REGION Network 7: LS425, LS442 Alarms (RIO 07: APT)
   RUNG wire#powerrail
      "1602_DIGITAL_HEALTH"(InputSignal := "20_TANKS_IP_DATA".RIO_07.FIRST_TANK.BWT_LEVEL_HIHI, InputTripLevel := #InputTripLevel, SensorHealthOut => "1092_HMI_OP_FLAGS".LS425_442_LevelSwitch_HighHigh_Alarm[14].Healthy, AlarmOut => "1092_HMI_OP_FLAGS".LS425_442_LevelSwitch_HighHigh_Alarm[14].UnhealthyAlarm)
   END_RUNG
   // the same network as SCL:
   "1602_DIGITAL_HEALTH"(InputSignal := "20_TANKS_IP_DATA".RIO_07.FIRST_TANK.BWT_LEVEL_HIHI,
                         InputTripLevel := #InputTripLevel,
                         SensorHealthOut => "1092_HMI_OP_FLAGS".LS425_442_LevelSwitch_HighHigh_Alarm[14].Healthy,
                         AlarmOut => "1092_HMI_OP_FLAGS".LS425_442_LevelSwitch_HighHigh_Alarm[14].UnhealthyAlarm);
END_REGION
END_FUNCTION

// folder: 1000 - 1999 BWT System Control/1060 - 1089 Alarm & Valve Status Handling/1080 - 1084 Tank Group Alarms

FUNCTION "1080_PT424_ALARMS" : Void   // FC1080, LAD
{ S7_Optimized_Access := 'TRUE' }
VERSION : 0.1
// Alarm wrapper function for Ullage Space Pressure Transmitter on each tank group.
BEGIN

REGION Network 1: PT424 Alarms (RIO 01)
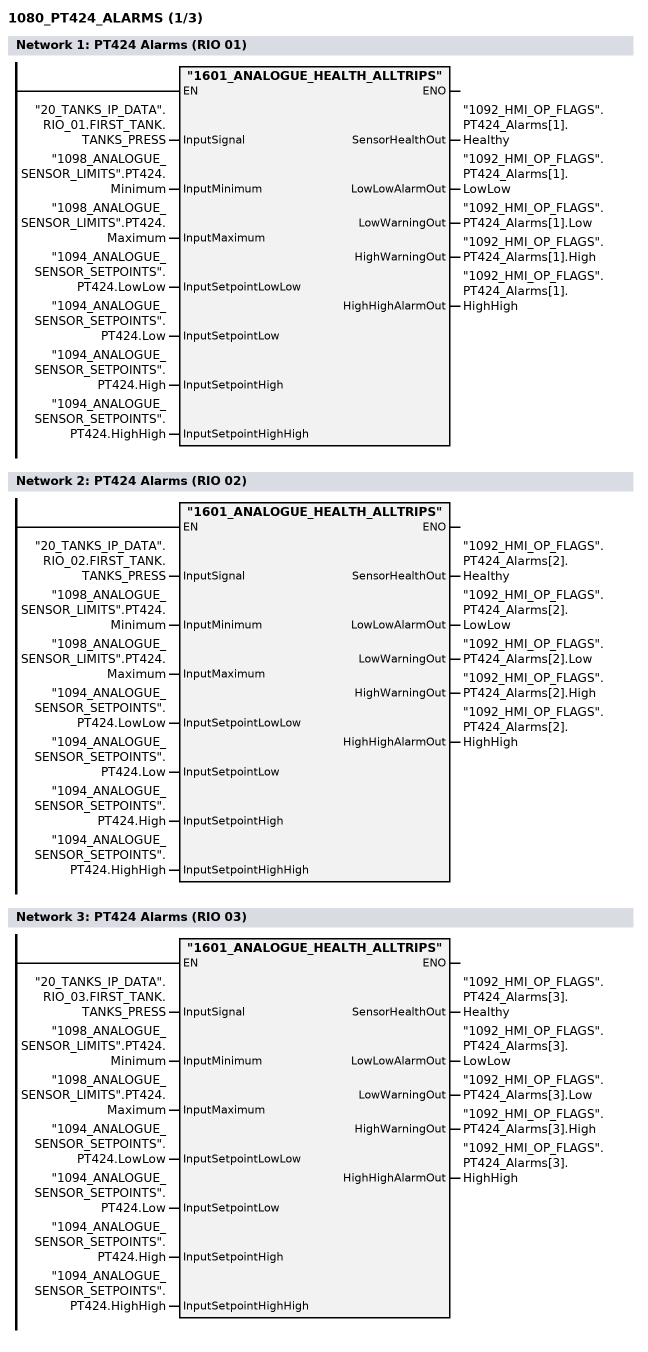
   RUNG wire#powerrail
      "1601_ANALOGUE_HEALTH_ALLTRIPS"(InputSignal := "20_TANKS_IP_DATA".RIO_01.FIRST_TANK.TANKS_PRESS, InputMinimum := "1098_ANALOGUE_SENSOR_LIMITS".PT424.Minimum, InputMaximum := "1098_ANALOGUE_SENSOR_LIMITS".PT424.Maximum, InputSetpointLowLow := "1094_ANALOGUE_SENSOR_SETPOINTS".PT424.LowLow, InputSetpointLow := "1094_ANALOGUE_SENSOR_SETPOINTS".PT424.Low, InputSetpointHigh := "1094_ANALOGUE_SENSOR_SETPOINTS".PT424.High, InputSetpointHighHigh := "1094_ANALOGUE_SENSOR_SETPOINTS".PT424.HighHigh, SensorHealthOut => "1092_HMI_OP_FLAGS".PT424_Alarms[1].Healthy, LowLowAlarmOut => "1092_HMI_OP_FLAGS".PT424_Alarms[1].LowLow, LowWarningOut => "1092_HMI_OP_FLAGS".PT424_Alarms[1].Low, HighWarningOut => "1092_HMI_OP_FLAGS".PT424_Alarms[1].High, HighHighAlarmOut => "1092_HMI_OP_FLAGS".PT424_Alarms[1].HighHigh)
   END_RUNG
   // the same network as SCL:
   "1601_ANALOGUE_HEALTH_ALLTRIPS"(InputSignal := "20_TANKS_IP_DATA".RIO_01.FIRST_TANK.TANKS_PRESS,
                           InputMinimum := "1098_ANALOGUE_SENSOR_LIMITS".PT424.Minimum,
                           InputMaximum := "1098_ANALOGUE_SENSOR_LIMITS".PT424.Maximum,
                           InputSetpointLowLow := "1094_ANALOGUE_SENSOR_SETPOINTS".PT424.LowLow,
                           InputSetpointLow := "1094_ANALOGUE_SENSOR_SETPOINTS".PT424.Low,
                           InputSetpointHigh := "1094_ANALOGUE_SENSOR_SETPOINTS".PT424.High,
                           InputSetpointHighHigh := "1094_ANALOGUE_SENSOR_SETPOINTS".PT424.HighHigh,
                           SensorHealthOut => "1092_HMI_OP_FLAGS".PT424_Alarms[1].Healthy,
                           LowLowAlarmOut => "1092_HMI_OP_FLAGS".PT424_Alarms[1].LowLow,
                           LowWarningOut => "1092_HMI_OP_FLAGS".PT424_Alarms[1].Low,
                           HighWarningOut => "1092_HMI_OP_FLAGS".PT424_Alarms[1].High,
                           HighHighAlarmOut => "1092_HMI_OP_FLAGS".PT424_Alarms[1].HighHigh);
END_REGION

REGION Network 2: PT424 Alarms (RIO 02)
   RUNG wire#powerrail
      "1601_ANALOGUE_HEALTH_ALLTRIPS"(InputSignal := "20_TANKS_IP_DATA".RIO_02.FIRST_TANK.TANKS_PRESS, InputMinimum := "1098_ANALOGUE_SENSOR_LIMITS".PT424.Minimum, InputMaximum := "1098_ANALOGUE_SENSOR_LIMITS".PT424.Maximum, InputSetpointLowLow := "1094_ANALOGUE_SENSOR_SETPOINTS".PT424.LowLow, InputSetpointLow := "1094_ANALOGUE_SENSOR_SETPOINTS".PT424.Low, InputSetpointHigh := "1094_ANALOGUE_SENSOR_SETPOINTS".PT424.High, InputSetpointHighHigh := "1094_ANALOGUE_SENSOR_SETPOINTS".PT424.HighHigh, SensorHealthOut => "1092_HMI_OP_FLAGS".PT424_Alarms[2].Healthy, LowLowAlarmOut => "1092_HMI_OP_FLAGS".PT424_Alarms[2].LowLow, LowWarningOut => "1092_HMI_OP_FLAGS".PT424_Alarms[2].Low, HighWarningOut => "1092_HMI_OP_FLAGS".PT424_Alarms[2].High, HighHighAlarmOut => "1092_HMI_OP_FLAGS".PT424_Alarms[2].HighHigh)
   END_RUNG
   // the same network as SCL:
   "1601_ANALOGUE_HEALTH_ALLTRIPS"(InputSignal := "20_TANKS_IP_DATA".RIO_02.FIRST_TANK.TANKS_PRESS,
                           InputMinimum := "1098_ANALOGUE_SENSOR_LIMITS".PT424.Minimum,
                           InputMaximum := "1098_ANALOGUE_SENSOR_LIMITS".PT424.Maximum,
                           InputSetpointLowLow := "1094_ANALOGUE_SENSOR_SETPOINTS".PT424.LowLow,
                           InputSetpointLow := "1094_ANALOGUE_SENSOR_SETPOINTS".PT424.Low,
                           InputSetpointHigh := "1094_ANALOGUE_SENSOR_SETPOINTS".PT424.High,
                           InputSetpointHighHigh := "1094_ANALOGUE_SENSOR_SETPOINTS".PT424.HighHigh,
                           SensorHealthOut => "1092_HMI_OP_FLAGS".PT424_Alarms[2].Healthy,
                           LowLowAlarmOut => "1092_HMI_OP_FLAGS".PT424_Alarms[2].LowLow,
                           LowWarningOut => "1092_HMI_OP_FLAGS".PT424_Alarms[2].Low,
                           HighWarningOut => "1092_HMI_OP_FLAGS".PT424_Alarms[2].High,
                           HighHighAlarmOut => "1092_HMI_OP_FLAGS".PT424_Alarms[2].HighHigh);
END_REGION

REGION Network 3: PT424 Alarms (RIO 03)
   RUNG wire#powerrail
      "1601_ANALOGUE_HEALTH_ALLTRIPS"(InputSignal := "20_TANKS_IP_DATA".RIO_03.FIRST_TANK.TANKS_PRESS, InputMinimum := "1098_ANALOGUE_SENSOR_LIMITS".PT424.Minimum, InputMaximum := "1098_ANALOGUE_SENSOR_LIMITS".PT424.Maximum, InputSetpointLowLow := "1094_ANALOGUE_SENSOR_SETPOINTS".PT424.LowLow, InputSetpointLow := "1094_ANALOGUE_SENSOR_SETPOINTS".PT424.Low, InputSetpointHigh := "1094_ANALOGUE_SENSOR_SETPOINTS".PT424.High, InputSetpointHighHigh := "1094_ANALOGUE_SENSOR_SETPOINTS".PT424.HighHigh, SensorHealthOut => "1092_HMI_OP_FLAGS".PT424_Alarms[3].Healthy, LowLowAlarmOut => "1092_HMI_OP_FLAGS".PT424_Alarms[3].LowLow, LowWarningOut => "1092_HMI_OP_FLAGS".PT424_Alarms[3].Low, HighWarningOut => "1092_HMI_OP_FLAGS".PT424_Alarms[3].High, HighHighAlarmOut => "1092_HMI_OP_FLAGS".PT424_Alarms[3].HighHigh)
   END_RUNG
   // the same network as SCL:
   "1601_ANALOGUE_HEALTH_ALLTRIPS"(InputSignal := "20_TANKS_IP_DATA".RIO_03.FIRST_TANK.TANKS_PRESS,
                           InputMinimum := "1098_ANALOGUE_SENSOR_LIMITS".PT424.Minimum,
                           InputMaximum := "1098_ANALOGUE_SENSOR_LIMITS".PT424.Maximum,
                           InputSetpointLowLow := "1094_ANALOGUE_SENSOR_SETPOINTS".PT424.LowLow,
                           InputSetpointLow := "1094_ANALOGUE_SENSOR_SETPOINTS".PT424.Low,
                           InputSetpointHigh := "1094_ANALOGUE_SENSOR_SETPOINTS".PT424.High,
                           InputSetpointHighHigh := "1094_ANALOGUE_SENSOR_SETPOINTS".PT424.HighHigh,
                           SensorHealthOut => "1092_HMI_OP_FLAGS".PT424_Alarms[3].Healthy,
                           LowLowAlarmOut => "1092_HMI_OP_FLAGS".PT424_Alarms[3].LowLow,
                           LowWarningOut => "1092_HMI_OP_FLAGS".PT424_Alarms[3].Low,
                           HighWarningOut => "1092_HMI_OP_FLAGS".PT424_Alarms[3].High,
                           HighHighAlarmOut => "1092_HMI_OP_FLAGS".PT424_Alarms[3].HighHigh);
END_REGION

REGION Network 4: PT424 Alarms (RIO 04)
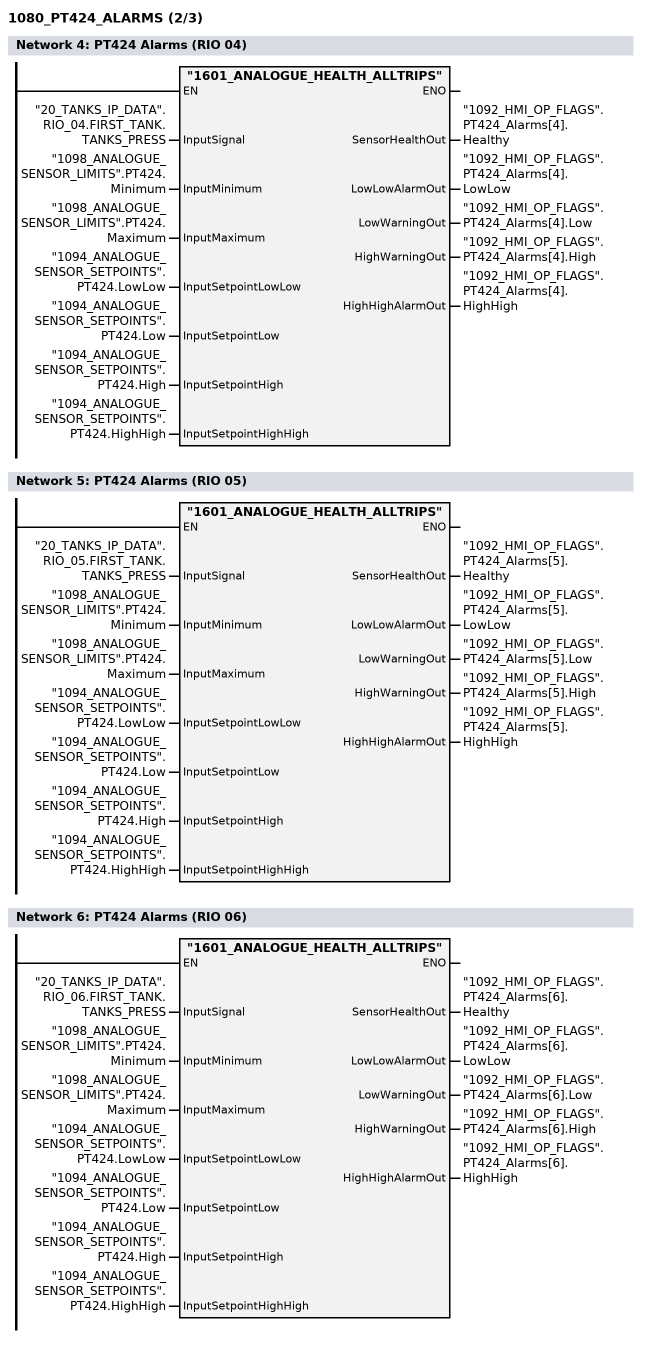
   RUNG wire#powerrail
      "1601_ANALOGUE_HEALTH_ALLTRIPS"(InputSignal := "20_TANKS_IP_DATA".RIO_04.FIRST_TANK.TANKS_PRESS, InputMinimum := "1098_ANALOGUE_SENSOR_LIMITS".PT424.Minimum, InputMaximum := "1098_ANALOGUE_SENSOR_LIMITS".PT424.Maximum, InputSetpointLowLow := "1094_ANALOGUE_SENSOR_SETPOINTS".PT424.LowLow, InputSetpointLow := "1094_ANALOGUE_SENSOR_SETPOINTS".PT424.Low, InputSetpointHigh := "1094_ANALOGUE_SENSOR_SETPOINTS".PT424.High, InputSetpointHighHigh := "1094_ANALOGUE_SENSOR_SETPOINTS".PT424.HighHigh, SensorHealthOut => "1092_HMI_OP_FLAGS".PT424_Alarms[4].Healthy, LowLowAlarmOut => "1092_HMI_OP_FLAGS".PT424_Alarms[4].LowLow, LowWarningOut => "1092_HMI_OP_FLAGS".PT424_Alarms[4].Low, HighWarningOut => "1092_HMI_OP_FLAGS".PT424_Alarms[4].High, HighHighAlarmOut => "1092_HMI_OP_FLAGS".PT424_Alarms[4].HighHigh)
   END_RUNG
   // the same network as SCL:
   "1601_ANALOGUE_HEALTH_ALLTRIPS"(InputSignal := "20_TANKS_IP_DATA".RIO_04.FIRST_TANK.TANKS_PRESS,
                           InputMinimum := "1098_ANALOGUE_SENSOR_LIMITS".PT424.Minimum,
                           InputMaximum := "1098_ANALOGUE_SENSOR_LIMITS".PT424.Maximum,
                           InputSetpointLowLow := "1094_ANALOGUE_SENSOR_SETPOINTS".PT424.LowLow,
                           InputSetpointLow := "1094_ANALOGUE_SENSOR_SETPOINTS".PT424.Low,
                           InputSetpointHigh := "1094_ANALOGUE_SENSOR_SETPOINTS".PT424.High,
                           InputSetpointHighHigh := "1094_ANALOGUE_SENSOR_SETPOINTS".PT424.HighHigh,
                           SensorHealthOut => "1092_HMI_OP_FLAGS".PT424_Alarms[4].Healthy,
                           LowLowAlarmOut => "1092_HMI_OP_FLAGS".PT424_Alarms[4].LowLow,
                           LowWarningOut => "1092_HMI_OP_FLAGS".PT424_Alarms[4].Low,
                           HighWarningOut => "1092_HMI_OP_FLAGS".PT424_Alarms[4].High,
                           HighHighAlarmOut => "1092_HMI_OP_FLAGS".PT424_Alarms[4].HighHigh);
END_REGION

REGION Network 5: PT424 Alarms (RIO 05)
   RUNG wire#powerrail
      "1601_ANALOGUE_HEALTH_ALLTRIPS"(InputSignal := "20_TANKS_IP_DATA".RIO_05.FIRST_TANK.TANKS_PRESS, InputMinimum := "1098_ANALOGUE_SENSOR_LIMITS".PT424.Minimum, InputMaximum := "1098_ANALOGUE_SENSOR_LIMITS".PT424.Maximum, InputSetpointLowLow := "1094_ANALOGUE_SENSOR_SETPOINTS".PT424.LowLow, InputSetpointLow := "1094_ANALOGUE_SENSOR_SETPOINTS".PT424.Low, InputSetpointHigh := "1094_ANALOGUE_SENSOR_SETPOINTS".PT424.High, InputSetpointHighHigh := "1094_ANALOGUE_SENSOR_SETPOINTS".PT424.HighHigh, SensorHealthOut => "1092_HMI_OP_FLAGS".PT424_Alarms[5].Healthy, LowLowAlarmOut => "1092_HMI_OP_FLAGS".PT424_Alarms[5].LowLow, LowWarningOut => "1092_HMI_OP_FLAGS".PT424_Alarms[5].Low, HighWarningOut => "1092_HMI_OP_FLAGS".PT424_Alarms[5].High, HighHighAlarmOut => "1092_HMI_OP_FLAGS".PT424_Alarms[5].HighHigh)
   END_RUNG
   // the same network as SCL:
   "1601_ANALOGUE_HEALTH_ALLTRIPS"(InputSignal := "20_TANKS_IP_DATA".RIO_05.FIRST_TANK.TANKS_PRESS,
                           InputMinimum := "1098_ANALOGUE_SENSOR_LIMITS".PT424.Minimum,
                           InputMaximum := "1098_ANALOGUE_SENSOR_LIMITS".PT424.Maximum,
                           InputSetpointLowLow := "1094_ANALOGUE_SENSOR_SETPOINTS".PT424.LowLow,
                           InputSetpointLow := "1094_ANALOGUE_SENSOR_SETPOINTS".PT424.Low,
                           InputSetpointHigh := "1094_ANALOGUE_SENSOR_SETPOINTS".PT424.High,
                           InputSetpointHighHigh := "1094_ANALOGUE_SENSOR_SETPOINTS".PT424.HighHigh,
                           SensorHealthOut => "1092_HMI_OP_FLAGS".PT424_Alarms[5].Healthy,
                           LowLowAlarmOut => "1092_HMI_OP_FLAGS".PT424_Alarms[5].LowLow,
                           LowWarningOut => "1092_HMI_OP_FLAGS".PT424_Alarms[5].Low,
                           HighWarningOut => "1092_HMI_OP_FLAGS".PT424_Alarms[5].High,
                           HighHighAlarmOut => "1092_HMI_OP_FLAGS".PT424_Alarms[5].HighHigh);
END_REGION

REGION Network 6: PT424 Alarms (RIO 06)
   RUNG wire#powerrail
      "1601_ANALOGUE_HEALTH_ALLTRIPS"(InputSignal := "20_TANKS_IP_DATA".RIO_06.FIRST_TANK.TANKS_PRESS, InputMinimum := "1098_ANALOGUE_SENSOR_LIMITS".PT424.Minimum, InputMaximum := "1098_ANALOGUE_SENSOR_LIMITS".PT424.Maximum, InputSetpointLowLow := "1094_ANALOGUE_SENSOR_SETPOINTS".PT424.LowLow, InputSetpointLow := "1094_ANALOGUE_SENSOR_SETPOINTS".PT424.Low, InputSetpointHigh := "1094_ANALOGUE_SENSOR_SETPOINTS".PT424.High, InputSetpointHighHigh := "1094_ANALOGUE_SENSOR_SETPOINTS".PT424.HighHigh, SensorHealthOut => "1092_HMI_OP_FLAGS".PT424_Alarms[6].Healthy, LowLowAlarmOut => "1092_HMI_OP_FLAGS".PT424_Alarms[6].LowLow, LowWarningOut => "1092_HMI_OP_FLAGS".PT424_Alarms[6].Low, HighWarningOut => "1092_HMI_OP_FLAGS".PT424_Alarms[6].High, HighHighAlarmOut => "1092_HMI_OP_FLAGS".PT424_Alarms[6].HighHigh)
   END_RUNG
   // the same network as SCL:
   "1601_ANALOGUE_HEALTH_ALLTRIPS"(InputSignal := "20_TANKS_IP_DATA".RIO_06.FIRST_TANK.TANKS_PRESS,
                           InputMinimum := "1098_ANALOGUE_SENSOR_LIMITS".PT424.Minimum,
                           InputMaximum := "1098_ANALOGUE_SENSOR_LIMITS".PT424.Maximum,
                           InputSetpointLowLow := "1094_ANALOGUE_SENSOR_SETPOINTS".PT424.LowLow,
                           InputSetpointLow := "1094_ANALOGUE_SENSOR_SETPOINTS".PT424.Low,
                           InputSetpointHigh := "1094_ANALOGUE_SENSOR_SETPOINTS".PT424.High,
                           InputSetpointHighHigh := "1094_ANALOGUE_SENSOR_SETPOINTS".PT424.HighHigh,
                           SensorHealthOut => "1092_HMI_OP_FLAGS".PT424_Alarms[6].Healthy,
                           LowLowAlarmOut => "1092_HMI_OP_FLAGS".PT424_Alarms[6].LowLow,
                           LowWarningOut => "1092_HMI_OP_FLAGS".PT424_Alarms[6].Low,
                           HighWarningOut => "1092_HMI_OP_FLAGS".PT424_Alarms[6].High,
                           HighHighAlarmOut => "1092_HMI_OP_FLAGS".PT424_Alarms[6].HighHigh);
END_REGION

REGION Network 7: PT424 Alarms (RIO 07)
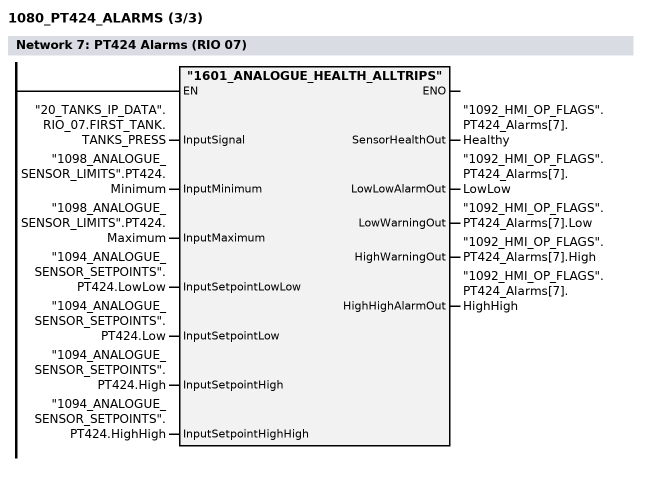
   RUNG wire#powerrail
      "1601_ANALOGUE_HEALTH_ALLTRIPS"(InputSignal := "20_TANKS_IP_DATA".RIO_07.FIRST_TANK.TANKS_PRESS, InputMinimum := "1098_ANALOGUE_SENSOR_LIMITS".PT424.Minimum, InputMaximum := "1098_ANALOGUE_SENSOR_LIMITS".PT424.Maximum, InputSetpointLowLow := "1094_ANALOGUE_SENSOR_SETPOINTS".PT424.LowLow, InputSetpointLow := "1094_ANALOGUE_SENSOR_SETPOINTS".PT424.Low, InputSetpointHigh := "1094_ANALOGUE_SENSOR_SETPOINTS".PT424.High, InputSetpointHighHigh := "1094_ANALOGUE_SENSOR_SETPOINTS".PT424.HighHigh, SensorHealthOut => "1092_HMI_OP_FLAGS".PT424_Alarms[7].Healthy, LowLowAlarmOut => "1092_HMI_OP_FLAGS".PT424_Alarms[7].LowLow, LowWarningOut => "1092_HMI_OP_FLAGS".PT424_Alarms[7].Low, HighWarningOut => "1092_HMI_OP_FLAGS".PT424_Alarms[7].High, HighHighAlarmOut => "1092_HMI_OP_FLAGS".PT424_Alarms[7].HighHigh)
   END_RUNG
   // the same network as SCL:
   "1601_ANALOGUE_HEALTH_ALLTRIPS"(InputSignal := "20_TANKS_IP_DATA".RIO_07.FIRST_TANK.TANKS_PRESS,
                           InputMinimum := "1098_ANALOGUE_SENSOR_LIMITS".PT424.Minimum,
                           InputMaximum := "1098_ANALOGUE_SENSOR_LIMITS".PT424.Maximum,
                           InputSetpointLowLow := "1094_ANALOGUE_SENSOR_SETPOINTS".PT424.LowLow,
                           InputSetpointLow := "1094_ANALOGUE_SENSOR_SETPOINTS".PT424.Low,
                           InputSetpointHigh := "1094_ANALOGUE_SENSOR_SETPOINTS".PT424.High,
                           InputSetpointHighHigh := "1094_ANALOGUE_SENSOR_SETPOINTS".PT424.HighHigh,
                           SensorHealthOut => "1092_HMI_OP_FLAGS".PT424_Alarms[7].Healthy,
                           LowLowAlarmOut => "1092_HMI_OP_FLAGS".PT424_Alarms[7].LowLow,
                           LowWarningOut => "1092_HMI_OP_FLAGS".PT424_Alarms[7].Low,
                           HighWarningOut => "1092_HMI_OP_FLAGS".PT424_Alarms[7].High,
                           HighHighAlarmOut => "1092_HMI_OP_FLAGS".PT424_Alarms[7].HighHigh);
END_REGION
END_FUNCTION

FUNCTION "1081_PS436_ALARMS" : Void   // FC1081, LAD
{ S7_Optimized_Access := 'TRUE' }
VERSION : 0.1
// Alarm wrapper function for Ullage Space Pressure Switch on each tank group.
   VAR CONSTANT
      InputTripLevel : Bool := true;   // The input trip level for this function, if the input is equal to this digital value, trip the alarm.
   END_VAR
BEGIN

REGION Network 1: PT424 Alarms (RIO 01)
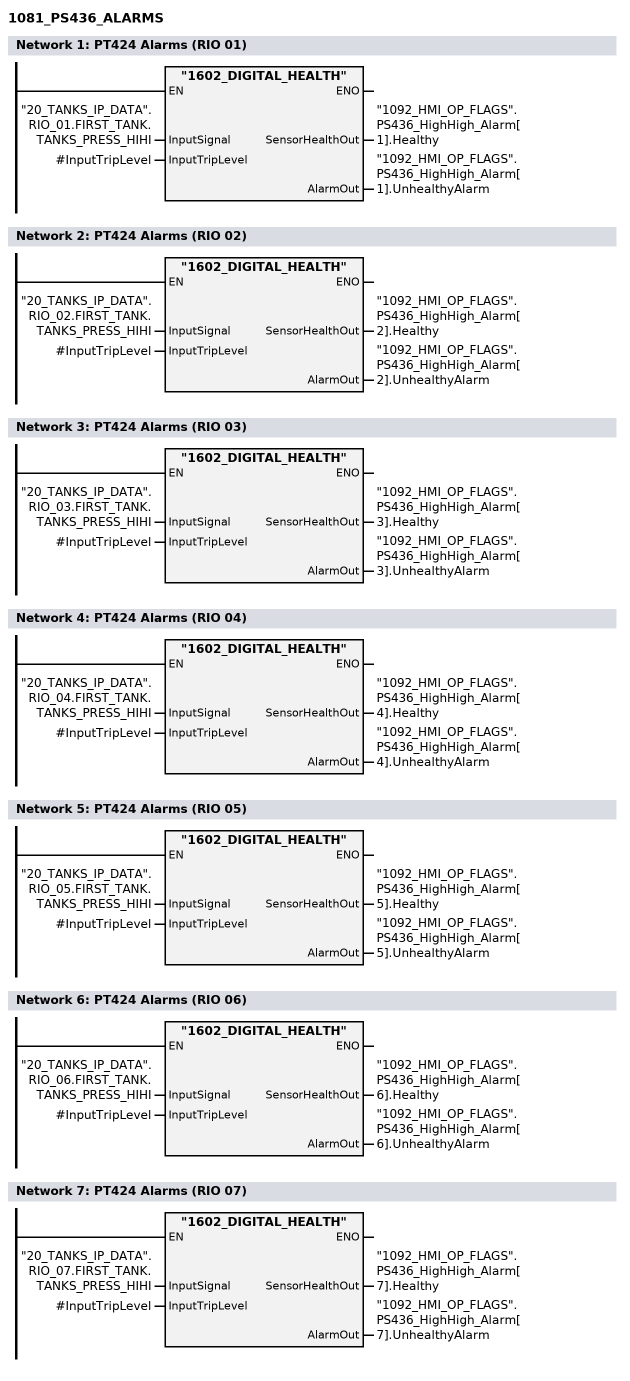
   RUNG wire#powerrail
      "1602_DIGITAL_HEALTH"(InputSignal := "20_TANKS_IP_DATA".RIO_01.FIRST_TANK.TANKS_PRESS_HIHI, InputTripLevel := #InputTripLevel, SensorHealthOut => "1092_HMI_OP_FLAGS".PS436_HighHigh_Alarm[1].Healthy, AlarmOut => "1092_HMI_OP_FLAGS".PS436_HighHigh_Alarm[1].UnhealthyAlarm)
   END_RUNG
   // the same network as SCL:
   "1602_DIGITAL_HEALTH"(InputSignal := "20_TANKS_IP_DATA".RIO_01.FIRST_TANK.TANKS_PRESS_HIHI,
                         InputTripLevel := #InputTripLevel,
                         SensorHealthOut => "1092_HMI_OP_FLAGS".PS436_HighHigh_Alarm[1].Healthy,
                         AlarmOut => "1092_HMI_OP_FLAGS".PS436_HighHigh_Alarm[1].UnhealthyAlarm);
END_REGION

REGION Network 2: PT424 Alarms (RIO 02)
   RUNG wire#powerrail
      "1602_DIGITAL_HEALTH"(InputSignal := "20_TANKS_IP_DATA".RIO_02.FIRST_TANK.TANKS_PRESS_HIHI, InputTripLevel := #InputTripLevel, SensorHealthOut => "1092_HMI_OP_FLAGS".PS436_HighHigh_Alarm[2].Healthy, AlarmOut => "1092_HMI_OP_FLAGS".PS436_HighHigh_Alarm[2].UnhealthyAlarm)
   END_RUNG
   // the same network as SCL:
   "1602_DIGITAL_HEALTH"(InputSignal := "20_TANKS_IP_DATA".RIO_02.FIRST_TANK.TANKS_PRESS_HIHI,
                         InputTripLevel := #InputTripLevel,
                         SensorHealthOut => "1092_HMI_OP_FLAGS".PS436_HighHigh_Alarm[2].Healthy,
                         AlarmOut => "1092_HMI_OP_FLAGS".PS436_HighHigh_Alarm[2].UnhealthyAlarm);
END_REGION

REGION Network 3: PT424 Alarms (RIO 03)
   RUNG wire#powerrail
      "1602_DIGITAL_HEALTH"(InputSignal := "20_TANKS_IP_DATA".RIO_03.FIRST_TANK.TANKS_PRESS_HIHI, InputTripLevel := #InputTripLevel, SensorHealthOut => "1092_HMI_OP_FLAGS".PS436_HighHigh_Alarm[3].Healthy, AlarmOut => "1092_HMI_OP_FLAGS".PS436_HighHigh_Alarm[3].UnhealthyAlarm)
   END_RUNG
   // the same network as SCL:
   "1602_DIGITAL_HEALTH"(InputSignal := "20_TANKS_IP_DATA".RIO_03.FIRST_TANK.TANKS_PRESS_HIHI,
                         InputTripLevel := #InputTripLevel,
                         SensorHealthOut => "1092_HMI_OP_FLAGS".PS436_HighHigh_Alarm[3].Healthy,
                         AlarmOut => "1092_HMI_OP_FLAGS".PS436_HighHigh_Alarm[3].UnhealthyAlarm);
END_REGION

REGION Network 4: PT424 Alarms (RIO 04)
   RUNG wire#powerrail
      "1602_DIGITAL_HEALTH"(InputSignal := "20_TANKS_IP_DATA".RIO_04.FIRST_TANK.TANKS_PRESS_HIHI, InputTripLevel := #InputTripLevel, SensorHealthOut => "1092_HMI_OP_FLAGS".PS436_HighHigh_Alarm[4].Healthy, AlarmOut => "1092_HMI_OP_FLAGS".PS436_HighHigh_Alarm[4].UnhealthyAlarm)
   END_RUNG
   // the same network as SCL:
   "1602_DIGITAL_HEALTH"(InputSignal := "20_TANKS_IP_DATA".RIO_04.FIRST_TANK.TANKS_PRESS_HIHI,
                         InputTripLevel := #InputTripLevel,
                         SensorHealthOut => "1092_HMI_OP_FLAGS".PS436_HighHigh_Alarm[4].Healthy,
                         AlarmOut => "1092_HMI_OP_FLAGS".PS436_HighHigh_Alarm[4].UnhealthyAlarm);
END_REGION

REGION Network 5: PT424 Alarms (RIO 05)
   RUNG wire#powerrail
      "1602_DIGITAL_HEALTH"(InputSignal := "20_TANKS_IP_DATA".RIO_05.FIRST_TANK.TANKS_PRESS_HIHI, InputTripLevel := #InputTripLevel, SensorHealthOut => "1092_HMI_OP_FLAGS".PS436_HighHigh_Alarm[5].Healthy, AlarmOut => "1092_HMI_OP_FLAGS".PS436_HighHigh_Alarm[5].UnhealthyAlarm)
   END_RUNG
   // the same network as SCL:
   "1602_DIGITAL_HEALTH"(InputSignal := "20_TANKS_IP_DATA".RIO_05.FIRST_TANK.TANKS_PRESS_HIHI,
                         InputTripLevel := #InputTripLevel,
                         SensorHealthOut => "1092_HMI_OP_FLAGS".PS436_HighHigh_Alarm[5].Healthy,
                         AlarmOut => "1092_HMI_OP_FLAGS".PS436_HighHigh_Alarm[5].UnhealthyAlarm);
END_REGION

REGION Network 6: PT424 Alarms (RIO 06)
   RUNG wire#powerrail
      "1602_DIGITAL_HEALTH"(InputSignal := "20_TANKS_IP_DATA".RIO_06.FIRST_TANK.TANKS_PRESS_HIHI, InputTripLevel := #InputTripLevel, SensorHealthOut => "1092_HMI_OP_FLAGS".PS436_HighHigh_Alarm[6].Healthy, AlarmOut => "1092_HMI_OP_FLAGS".PS436_HighHigh_Alarm[6].UnhealthyAlarm)
   END_RUNG
   // the same network as SCL:
   "1602_DIGITAL_HEALTH"(InputSignal := "20_TANKS_IP_DATA".RIO_06.FIRST_TANK.TANKS_PRESS_HIHI,
                         InputTripLevel := #InputTripLevel,
                         SensorHealthOut => "1092_HMI_OP_FLAGS".PS436_HighHigh_Alarm[6].Healthy,
                         AlarmOut => "1092_HMI_OP_FLAGS".PS436_HighHigh_Alarm[6].UnhealthyAlarm);
END_REGION

REGION Network 7: PT424 Alarms (RIO 07)
   RUNG wire#powerrail
      "1602_DIGITAL_HEALTH"(InputSignal := "20_TANKS_IP_DATA".RIO_07.FIRST_TANK.TANKS_PRESS_HIHI, InputTripLevel := #InputTripLevel, SensorHealthOut => "1092_HMI_OP_FLAGS".PS436_HighHigh_Alarm[7].Healthy, AlarmOut => "1092_HMI_OP_FLAGS".PS436_HighHigh_Alarm[7].UnhealthyAlarm)
   END_RUNG
   // the same network as SCL:
   "1602_DIGITAL_HEALTH"(InputSignal := "20_TANKS_IP_DATA".RIO_07.FIRST_TANK.TANKS_PRESS_HIHI,
                         InputTripLevel := #InputTripLevel,
                         SensorHealthOut => "1092_HMI_OP_FLAGS".PS436_HighHigh_Alarm[7].Healthy,
                         AlarmOut => "1092_HMI_OP_FLAGS".PS436_HighHigh_Alarm[7].UnhealthyAlarm);
END_REGION
END_FUNCTION

// folder: 1000 - 1999 BWT System Control/1060 - 1089 Alarm & Valve Status Handling/1085 - 1090 Valve Statuses

FUNCTION "1085_600CV421_422_STATUS" : Void   // FC1085, LAD
{ S7_Optimized_Access := 'TRUE' }
VERSION : 0.1
// Calculate the valve status' for each of the Gas To Tank Inlet Valves.
BEGIN

REGION Network 1: 600-CV-421, 600-CV-422 Alarms (RIO 01: FPT. 1P, 1S)
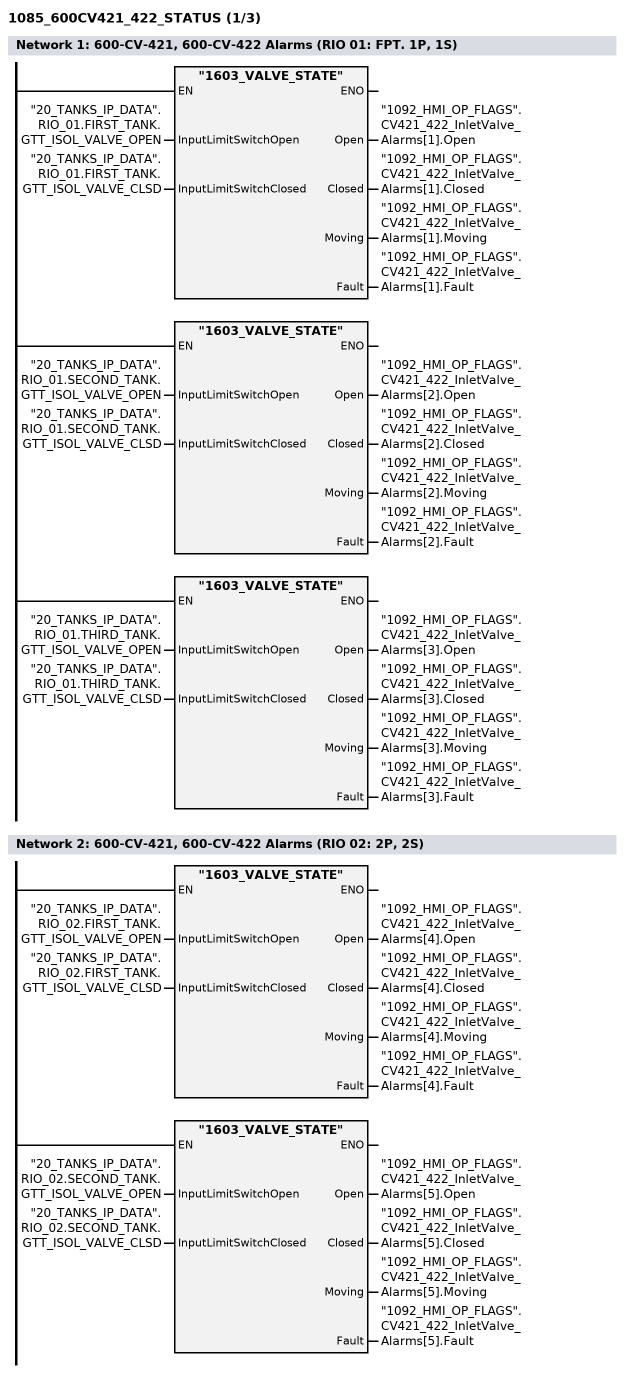
   RUNG wire#powerrail
      "1603_VALVE_STATE"(InputLimitSwitchOpen := "20_TANKS_IP_DATA".RIO_01.FIRST_TANK.GTT_ISOL_VALVE_OPEN, InputLimitSwitchClosed := "20_TANKS_IP_DATA".RIO_01.FIRST_TANK.GTT_ISOL_VALVE_CLSD, Open => "1092_HMI_OP_FLAGS".CV421_422_InletValve_Alarms[1].Open, Closed => "1092_HMI_OP_FLAGS".CV421_422_InletValve_Alarms[1].Closed, Moving => "1092_HMI_OP_FLAGS".CV421_422_InletValve_Alarms[1].Moving, Fault => "1092_HMI_OP_FLAGS".CV421_422_InletValve_Alarms[1].Fault)
   END_RUNG
   RUNG wire#powerrail
      "1603_VALVE_STATE"(InputLimitSwitchOpen := "20_TANKS_IP_DATA".RIO_01.SECOND_TANK.GTT_ISOL_VALVE_OPEN, InputLimitSwitchClosed := "20_TANKS_IP_DATA".RIO_01.SECOND_TANK.GTT_ISOL_VALVE_CLSD, Open => "1092_HMI_OP_FLAGS".CV421_422_InletValve_Alarms[2].Open, Closed => "1092_HMI_OP_FLAGS".CV421_422_InletValve_Alarms[2].Closed, Moving => "1092_HMI_OP_FLAGS".CV421_422_InletValve_Alarms[2].Moving, Fault => "1092_HMI_OP_FLAGS".CV421_422_InletValve_Alarms[2].Fault)
   END_RUNG
   RUNG wire#powerrail
      "1603_VALVE_STATE"(InputLimitSwitchOpen := "20_TANKS_IP_DATA".RIO_01.THIRD_TANK.GTT_ISOL_VALVE_OPEN, InputLimitSwitchClosed := "20_TANKS_IP_DATA".RIO_01.THIRD_TANK.GTT_ISOL_VALVE_CLSD, Open => "1092_HMI_OP_FLAGS".CV421_422_InletValve_Alarms[3].Open, Closed => "1092_HMI_OP_FLAGS".CV421_422_InletValve_Alarms[3].Closed, Moving => "1092_HMI_OP_FLAGS".CV421_422_InletValve_Alarms[3].Moving, Fault => "1092_HMI_OP_FLAGS".CV421_422_InletValve_Alarms[3].Fault)
   END_RUNG
   // the same network as SCL:
   "1603_VALVE_STATE"(InputLimitSwitchOpen := "20_TANKS_IP_DATA".RIO_01.FIRST_TANK.GTT_ISOL_VALVE_OPEN,
                      InputLimitSwitchClosed := "20_TANKS_IP_DATA".RIO_01.FIRST_TANK.GTT_ISOL_VALVE_CLSD,
                      Open => "1092_HMI_OP_FLAGS".CV421_422_InletValve_Alarms[1].Open,
                      Closed => "1092_HMI_OP_FLAGS".CV421_422_InletValve_Alarms[1].Closed,
                      Moving => "1092_HMI_OP_FLAGS".CV421_422_InletValve_Alarms[1].Moving,
                      Fault => "1092_HMI_OP_FLAGS".CV421_422_InletValve_Alarms[1].Fault);
   "1603_VALVE_STATE"(InputLimitSwitchOpen := "20_TANKS_IP_DATA".RIO_01.SECOND_TANK.GTT_ISOL_VALVE_OPEN,
                      InputLimitSwitchClosed := "20_TANKS_IP_DATA".RIO_01.SECOND_TANK.GTT_ISOL_VALVE_CLSD,
                      Open => "1092_HMI_OP_FLAGS".CV421_422_InletValve_Alarms[2].Open,
                      Closed => "1092_HMI_OP_FLAGS".CV421_422_InletValve_Alarms[2].Closed,
                      Moving => "1092_HMI_OP_FLAGS".CV421_422_InletValve_Alarms[2].Moving,
                      Fault => "1092_HMI_OP_FLAGS".CV421_422_InletValve_Alarms[2].Fault);
   "1603_VALVE_STATE"(InputLimitSwitchOpen := "20_TANKS_IP_DATA".RIO_01.THIRD_TANK.GTT_ISOL_VALVE_OPEN,
                      InputLimitSwitchClosed := "20_TANKS_IP_DATA".RIO_01.THIRD_TANK.GTT_ISOL_VALVE_CLSD,
                      Open => "1092_HMI_OP_FLAGS".CV421_422_InletValve_Alarms[3].Open,
                      Closed => "1092_HMI_OP_FLAGS".CV421_422_InletValve_Alarms[3].Closed,
                      Moving => "1092_HMI_OP_FLAGS".CV421_422_InletValve_Alarms[3].Moving,
                      Fault => "1092_HMI_OP_FLAGS".CV421_422_InletValve_Alarms[3].Fault);
END_REGION

REGION Network 2: 600-CV-421, 600-CV-422 Alarms (RIO 02: 2P, 2S)
   RUNG wire#powerrail
      "1603_VALVE_STATE"(InputLimitSwitchOpen := "20_TANKS_IP_DATA".RIO_02.FIRST_TANK.GTT_ISOL_VALVE_OPEN, InputLimitSwitchClosed := "20_TANKS_IP_DATA".RIO_02.FIRST_TANK.GTT_ISOL_VALVE_CLSD, Open => "1092_HMI_OP_FLAGS".CV421_422_InletValve_Alarms[4].Open, Closed => "1092_HMI_OP_FLAGS".CV421_422_InletValve_Alarms[4].Closed, Moving => "1092_HMI_OP_FLAGS".CV421_422_InletValve_Alarms[4].Moving, Fault => "1092_HMI_OP_FLAGS".CV421_422_InletValve_Alarms[4].Fault)
   END_RUNG
   RUNG wire#powerrail
      "1603_VALVE_STATE"(InputLimitSwitchOpen := "20_TANKS_IP_DATA".RIO_02.SECOND_TANK.GTT_ISOL_VALVE_OPEN, InputLimitSwitchClosed := "20_TANKS_IP_DATA".RIO_02.SECOND_TANK.GTT_ISOL_VALVE_CLSD, Open => "1092_HMI_OP_FLAGS".CV421_422_InletValve_Alarms[5].Open, Closed => "1092_HMI_OP_FLAGS".CV421_422_InletValve_Alarms[5].Closed, Moving => "1092_HMI_OP_FLAGS".CV421_422_InletValve_Alarms[5].Moving, Fault => "1092_HMI_OP_FLAGS".CV421_422_InletValve_Alarms[5].Fault)
   END_RUNG
   // the same network as SCL:
   "1603_VALVE_STATE"(InputLimitSwitchOpen := "20_TANKS_IP_DATA".RIO_02.FIRST_TANK.GTT_ISOL_VALVE_OPEN,
                      InputLimitSwitchClosed := "20_TANKS_IP_DATA".RIO_02.FIRST_TANK.GTT_ISOL_VALVE_CLSD,
                      Open => "1092_HMI_OP_FLAGS".CV421_422_InletValve_Alarms[4].Open,
                      Closed => "1092_HMI_OP_FLAGS".CV421_422_InletValve_Alarms[4].Closed,
                      Moving => "1092_HMI_OP_FLAGS".CV421_422_InletValve_Alarms[4].Moving,
                      Fault => "1092_HMI_OP_FLAGS".CV421_422_InletValve_Alarms[4].Fault);
   "1603_VALVE_STATE"(InputLimitSwitchOpen := "20_TANKS_IP_DATA".RIO_02.SECOND_TANK.GTT_ISOL_VALVE_OPEN,
                      InputLimitSwitchClosed := "20_TANKS_IP_DATA".RIO_02.SECOND_TANK.GTT_ISOL_VALVE_CLSD,
                      Open => "1092_HMI_OP_FLAGS".CV421_422_InletValve_Alarms[5].Open,
                      Closed => "1092_HMI_OP_FLAGS".CV421_422_InletValve_Alarms[5].Closed,
                      Moving => "1092_HMI_OP_FLAGS".CV421_422_InletValve_Alarms[5].Moving,
                      Fault => "1092_HMI_OP_FLAGS".CV421_422_InletValve_Alarms[5].Fault);
END_REGION

REGION Network 3: 600-CV-421, 600-CV-422 Alarms (RIO 03: 3P, 3S)
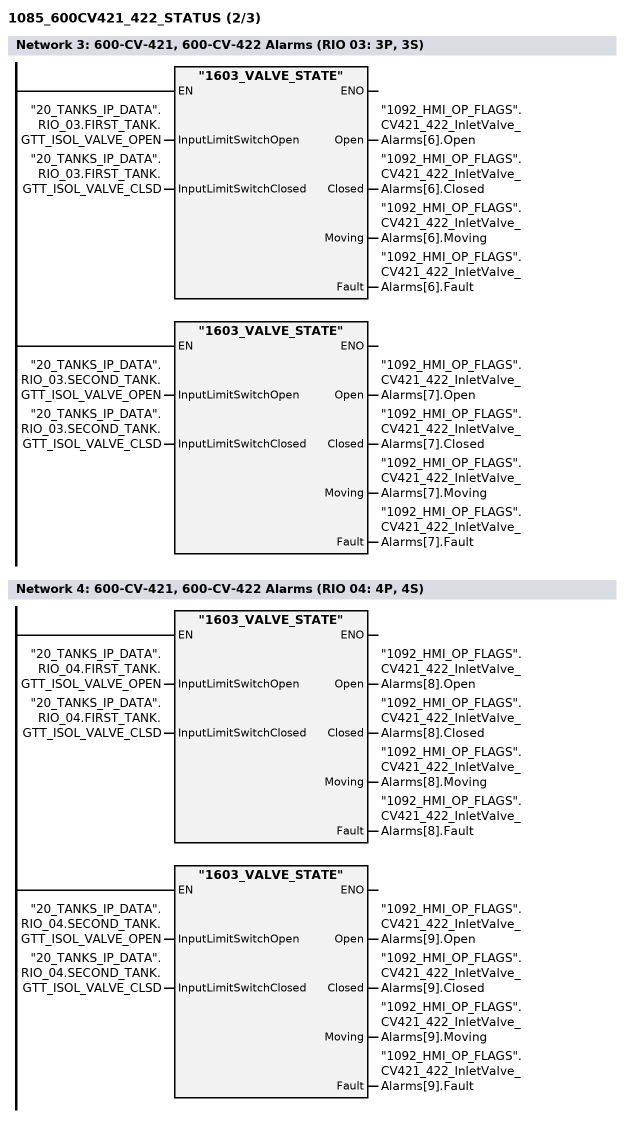
   RUNG wire#powerrail
      "1603_VALVE_STATE"(InputLimitSwitchOpen := "20_TANKS_IP_DATA".RIO_03.FIRST_TANK.GTT_ISOL_VALVE_OPEN, InputLimitSwitchClosed := "20_TANKS_IP_DATA".RIO_03.FIRST_TANK.GTT_ISOL_VALVE_CLSD, Open => "1092_HMI_OP_FLAGS".CV421_422_InletValve_Alarms[6].Open, Closed => "1092_HMI_OP_FLAGS".CV421_422_InletValve_Alarms[6].Closed, Moving => "1092_HMI_OP_FLAGS".CV421_422_InletValve_Alarms[6].Moving, Fault => "1092_HMI_OP_FLAGS".CV421_422_InletValve_Alarms[6].Fault)
   END_RUNG
   RUNG wire#powerrail
      "1603_VALVE_STATE"(InputLimitSwitchOpen := "20_TANKS_IP_DATA".RIO_03.SECOND_TANK.GTT_ISOL_VALVE_OPEN, InputLimitSwitchClosed := "20_TANKS_IP_DATA".RIO_03.SECOND_TANK.GTT_ISOL_VALVE_CLSD, Open => "1092_HMI_OP_FLAGS".CV421_422_InletValve_Alarms[7].Open, Closed => "1092_HMI_OP_FLAGS".CV421_422_InletValve_Alarms[7].Closed, Moving => "1092_HMI_OP_FLAGS".CV421_422_InletValve_Alarms[7].Moving, Fault => "1092_HMI_OP_FLAGS".CV421_422_InletValve_Alarms[7].Fault)
   END_RUNG
   // the same network as SCL:
   "1603_VALVE_STATE"(InputLimitSwitchOpen := "20_TANKS_IP_DATA".RIO_03.FIRST_TANK.GTT_ISOL_VALVE_OPEN,
                      InputLimitSwitchClosed := "20_TANKS_IP_DATA".RIO_03.FIRST_TANK.GTT_ISOL_VALVE_CLSD,
                      Open => "1092_HMI_OP_FLAGS".CV421_422_InletValve_Alarms[6].Open,
                      Closed => "1092_HMI_OP_FLAGS".CV421_422_InletValve_Alarms[6].Closed,
                      Moving => "1092_HMI_OP_FLAGS".CV421_422_InletValve_Alarms[6].Moving,
                      Fault => "1092_HMI_OP_FLAGS".CV421_422_InletValve_Alarms[6].Fault);
   "1603_VALVE_STATE"(InputLimitSwitchOpen := "20_TANKS_IP_DATA".RIO_03.SECOND_TANK.GTT_ISOL_VALVE_OPEN,
                      InputLimitSwitchClosed := "20_TANKS_IP_DATA".RIO_03.SECOND_TANK.GTT_ISOL_VALVE_CLSD,
                      Open => "1092_HMI_OP_FLAGS".CV421_422_InletValve_Alarms[7].Open,
                      Closed => "1092_HMI_OP_FLAGS".CV421_422_InletValve_Alarms[7].Closed,
                      Moving => "1092_HMI_OP_FLAGS".CV421_422_InletValve_Alarms[7].Moving,
                      Fault => "1092_HMI_OP_FLAGS".CV421_422_InletValve_Alarms[7].Fault);
END_REGION

REGION Network 4: 600-CV-421, 600-CV-422 Alarms (RIO 04: 4P, 4S)
   RUNG wire#powerrail
      "1603_VALVE_STATE"(InputLimitSwitchOpen := "20_TANKS_IP_DATA".RIO_04.FIRST_TANK.GTT_ISOL_VALVE_OPEN, InputLimitSwitchClosed := "20_TANKS_IP_DATA".RIO_04.FIRST_TANK.GTT_ISOL_VALVE_CLSD, Open => "1092_HMI_OP_FLAGS".CV421_422_InletValve_Alarms[8].Open, Closed => "1092_HMI_OP_FLAGS".CV421_422_InletValve_Alarms[8].Closed, Moving => "1092_HMI_OP_FLAGS".CV421_422_InletValve_Alarms[8].Moving, Fault => "1092_HMI_OP_FLAGS".CV421_422_InletValve_Alarms[8].Fault)
   END_RUNG
   RUNG wire#powerrail
      "1603_VALVE_STATE"(InputLimitSwitchOpen := "20_TANKS_IP_DATA".RIO_04.SECOND_TANK.GTT_ISOL_VALVE_OPEN, InputLimitSwitchClosed := "20_TANKS_IP_DATA".RIO_04.SECOND_TANK.GTT_ISOL_VALVE_CLSD, Open => "1092_HMI_OP_FLAGS".CV421_422_InletValve_Alarms[9].Open, Closed => "1092_HMI_OP_FLAGS".CV421_422_InletValve_Alarms[9].Closed, Moving => "1092_HMI_OP_FLAGS".CV421_422_InletValve_Alarms[9].Moving, Fault => "1092_HMI_OP_FLAGS".CV421_422_InletValve_Alarms[9].Fault)
   END_RUNG
   // the same network as SCL:
   "1603_VALVE_STATE"(InputLimitSwitchOpen := "20_TANKS_IP_DATA".RIO_04.FIRST_TANK.GTT_ISOL_VALVE_OPEN,
                      InputLimitSwitchClosed := "20_TANKS_IP_DATA".RIO_04.FIRST_TANK.GTT_ISOL_VALVE_CLSD,
                      Open => "1092_HMI_OP_FLAGS".CV421_422_InletValve_Alarms[8].Open,
                      Closed => "1092_HMI_OP_FLAGS".CV421_422_InletValve_Alarms[8].Closed,
                      Moving => "1092_HMI_OP_FLAGS".CV421_422_InletValve_Alarms[8].Moving,
                      Fault => "1092_HMI_OP_FLAGS".CV421_422_InletValve_Alarms[8].Fault);
   "1603_VALVE_STATE"(InputLimitSwitchOpen := "20_TANKS_IP_DATA".RIO_04.SECOND_TANK.GTT_ISOL_VALVE_OPEN,
                      InputLimitSwitchClosed := "20_TANKS_IP_DATA".RIO_04.SECOND_TANK.GTT_ISOL_VALVE_CLSD,
                      Open => "1092_HMI_OP_FLAGS".CV421_422_InletValve_Alarms[9].Open,
                      Closed => "1092_HMI_OP_FLAGS".CV421_422_InletValve_Alarms[9].Closed,
                      Moving => "1092_HMI_OP_FLAGS".CV421_422_InletValve_Alarms[9].Moving,
                      Fault => "1092_HMI_OP_FLAGS".CV421_422_InletValve_Alarms[9].Fault);
END_REGION

REGION Network 5: 600-CV-421, 600-CV-422 Alarms (RIO 05: 5P, 5S)